
   //-------------HEAD #5 PARAMETERS--------------------------

   "PLANT_CONSTANTS".CONST_rgtHeadPar[4].dParametersToDownload := 17;

   //Parameter IOfunct_LIO1
   "PLANT_CONSTANTS".CONST_rgtHeadPar[4].rgtAxisParameters[0].iAddress := 1826;
   "PLANT_CONSTANTS".CONST_rgtHeadPar[4].rgtAxisParameters[0].iLength := 2;
   "PLANT_CONSTANTS".CONST_rgtHeadPar[4].rgtAxisParameters[0].dValue := 20;

   //Parameter IOfunct_LIO2
   "PLANT_CONSTANTS".CONST_rgtHeadPar[4].rgtAxisParameters[1].iAddress := 1828;
   "PLANT_CONSTANTS".CONST_rgtHeadPar[4].rgtAxisParameters[1].iLength := 2;
   "PLANT_CONSTANTS".CONST_rgtHeadPar[4].rgtAxisParameters[1].dValue := 1;

   //Parameter IOfunct_LIO3
   "PLANT_CONSTANTS".CONST_rgtHeadPar[4].rgtAxisParameters[2].iAddress := 1830;
   "PLANT_CONSTANTS".CONST_rgtHeadPar[4].rgtAxisParameters[2].iLength := 2;
   "PLANT_CONSTANTS".CONST_rgtHeadPar[4].rgtAxisParameters[2].dValue := 1;

   //Parameter IOfunct_LIO4
   "PLANT_CONSTANTS".CONST_rgtHeadPar[4].rgtAxisParameters[3].iAddress := 1832;
   "PLANT_CONSTANTS".CONST_rgtHeadPar[4].rgtAxisParameters[3].iLength := 2;
   "PLANT_CONSTANTS".CONST_rgtHeadPar[4].rgtAxisParameters[3].dValue := 1;

   //Parameter IOsigLimN
   "PLANT_CONSTANTS".CONST_rgtHeadPar[4].rgtAxisParameters[4].iAddress := 1566;
   "PLANT_CONSTANTS".CONST_rgtHeadPar[4].rgtAxisParameters[4].iLength := 2;
   "PLANT_CONSTANTS".CONST_rgtHeadPar[4].rgtAxisParameters[4].dValue := 0;

   //Parameter IOsigLimP
   "PLANT_CONSTANTS".CONST_rgtHeadPar[4].rgtAxisParameters[5].iAddress := 1568;
   "PLANT_CONSTANTS".CONST_rgtHeadPar[4].rgtAxisParameters[5].iLength := 2;
   "PLANT_CONSTANTS".CONST_rgtHeadPar[4].rgtAxisParameters[5].dValue := 0;

   //Parameter IOsigRef
   "PLANT_CONSTANTS".CONST_rgtHeadPar[4].rgtAxisParameters[6].iAddress := 1564;
   "PLANT_CONSTANTS".CONST_rgtHeadPar[4].rgtAxisParameters[6].iLength := 2;
   "PLANT_CONSTANTS".CONST_rgtHeadPar[4].rgtAxisParameters[6].dValue := 2;

   //Parameter POSdirOfRotat
   "PLANT_CONSTANTS".CONST_rgtHeadPar[4].rgtAxisParameters[7].iAddress := 1560;
   "PLANT_CONSTANTS".CONST_rgtHeadPar[4].rgtAxisParameters[7].iLength := 2;
   "PLANT_CONSTANTS".CONST_rgtHeadPar[4].rgtAxisParameters[7].dValue := 0;

   //Parameter POSscaleDenom
   "PLANT_CONSTANTS".CONST_rgtHeadPar[4].rgtAxisParameters[8].iAddress := 1550;
   "PLANT_CONSTANTS".CONST_rgtHeadPar[4].rgtAxisParameters[8].iLength := 4;
   "PLANT_CONSTANTS".CONST_rgtHeadPar[4].rgtAxisParameters[8].dValue := 500;

   //Parameter POSscaleNum
   "PLANT_CONSTANTS".CONST_rgtHeadPar[4].rgtAxisParameters[9].iAddress := 1552;
   "PLANT_CONSTANTS".CONST_rgtHeadPar[4].rgtAxisParameters[9].iLength := 4;
   "PLANT_CONSTANTS".CONST_rgtHeadPar[4].rgtAxisParameters[9].dValue := 1;

   //Parameter RAMPacc
   "PLANT_CONSTANTS".CONST_rgtHeadPar[4].rgtAxisParameters[10].iAddress := 1556;
   "PLANT_CONSTANTS".CONST_rgtHeadPar[4].rgtAxisParameters[10].iLength := 4;
   "PLANT_CONSTANTS".CONST_rgtHeadPar[4].rgtAxisParameters[10].dValue := 20000;//[rot/s2]

   //Parameter RAMPdecel
   "PLANT_CONSTANTS".CONST_rgtHeadPar[4].rgtAxisParameters[11].iAddress := 1558;
   "PLANT_CONSTANTS".CONST_rgtHeadPar[4].rgtAxisParameters[11].iLength := 4;
   "PLANT_CONSTANTS".CONST_rgtHeadPar[4].rgtAxisParameters[11].dValue := 20000;//[rot/s2]

   //Parameter JOGn_fast
   "PLANT_CONSTANTS".CONST_rgtHeadPar[4].rgtAxisParameters[12].iAddress := 10506;
   "PLANT_CONSTANTS".CONST_rgtHeadPar[4].rgtAxisParameters[12].iLength := 2;
   "PLANT_CONSTANTS".CONST_rgtHeadPar[4].rgtAxisParameters[12].dValue := 1000;//[rot/min]

   //Parameter JOGn_slow
   "PLANT_CONSTANTS".CONST_rgtHeadPar[4].rgtAxisParameters[13].iAddress := 10504;
   "PLANT_CONSTANTS".CONST_rgtHeadPar[4].rgtAxisParameters[13].iLength := 2;
   "PLANT_CONSTANTS".CONST_rgtHeadPar[4].rgtAxisParameters[13].dValue := 1000;//[rot/min]

   //Parameter JOGstepusr
   "PLANT_CONSTANTS".CONST_rgtHeadPar[4].rgtAxisParameters[14].iAddress := 10510;
   "PLANT_CONSTANTS".CONST_rgtHeadPar[4].rgtAxisParameters[14].iLength := 4;
   "PLANT_CONSTANTS".CONST_rgtHeadPar[4].rgtAxisParameters[14].dValue := 0;

   //Parameter JOGtime
   "PLANT_CONSTANTS".CONST_rgtHeadPar[4].rgtAxisParameters[15].iAddress := 10512;
   "PLANT_CONSTANTS".CONST_rgtHeadPar[4].rgtAxisParameters[15].iLength := 2;
   "PLANT_CONSTANTS".CONST_rgtHeadPar[4].rgtAxisParameters[15].dValue := 1;

   //Parameter PAReeprSave ---MUST BE THE LAST!!!
   "PLANT_CONSTANTS".CONST_rgtHeadPar[4].rgtAxisParameters[16].iAddress := 1026;
   "PLANT_CONSTANTS".CONST_rgtHeadPar[4].rgtAxisParameters[16].iLength := 2;
   "PLANT_CONSTANTS".CONST_rgtHeadPar[4].rgtAxisParameters[16].dValue := 1;


   //-------------HEAD #6 PARAMETERS--------------------------

   "PLANT_CONSTANTS".CONST_rgtHeadPar[5].dParametersToDownload := 17;

   //Parameter IOfunct_LIO1
   "PLANT_CONSTANTS".CONST_rgtHeadPar[5].rgtAxisParameters[0].iAddress := 1826;
   "PLANT_CONSTANTS".CONST_rgtHeadPar[5].rgtAxisParameters[0].iLength := 2;
   "PLANT_CONSTANTS".CONST_rgtHeadPar[5].rgtAxisParameters[0].dValue := 20;

   //Parameter IOfunct_LIO2
   "PLANT_CONSTANTS".CONST_rgtHeadPar[5].rgtAxisParameters[1].iAddress := 1828;
   "PLANT_CONSTANTS".CONST_rgtHeadPar[5].rgtAxisParameters[1].iLength := 2;
   "PLANT_CONSTANTS".CONST_rgtHeadPar[5].rgtAxisParameters[1].dValue := 1;

   //Parameter IOfunct_LIO3
   "PLANT_CONSTANTS".CONST_rgtHeadPar[5].rgtAxisParameters[2].iAddress := 1830;
   "PLANT_CONSTANTS".CONST_rgtHeadPar[5].rgtAxisParameters[2].iLength := 2;
   "PLANT_CONSTANTS".CONST_rgtHeadPar[5].rgtAxisParameters[2].dValue := 1;

   //Parameter IOfunct_LIO4
   "PLANT_CONSTANTS".CONST_rgtHeadPar[5].rgtAxisParameters[3].iAddress := 1832;
   "PLANT_CONSTANTS".CONST_rgtHeadPar[5].rgtAxisParameters[3].iLength := 2;
   "PLANT_CONSTANTS".CONST_rgtHeadPar[5].rgtAxisParameters[3].dValue := 1;

   //Parameter IOsigLimN
   "PLANT_CONSTANTS".CONST_rgtHeadPar[5].rgtAxisParameters[4].iAddress := 1566;
   "PLANT_CONSTANTS".CONST_rgtHeadPar[5].rgtAxisParameters[4].iLength := 2;
   "PLANT_CONSTANTS".CONST_rgtHeadPar[5].rgtAxisParameters[4].dValue := 0;

   //Parameter IOsigLimP
   "PLANT_CONSTANTS".CONST_rgtHeadPar[5].rgtAxisParameters[5].iAddress := 1568;
   "PLANT_CONSTANTS".CONST_rgtHeadPar[5].rgtAxisParameters[5].iLength := 2;
   "PLANT_CONSTANTS".CONST_rgtHeadPar[5].rgtAxisParameters[5].dValue := 0;

   //Parameter IOsigRef
   "PLANT_CONSTANTS".CONST_rgtHeadPar[5].rgtAxisParameters[6].iAddress := 1564;
   "PLANT_CONSTANTS".CONST_rgtHeadPar[5].rgtAxisParameters[6].iLength := 2;
   "PLANT_CONSTANTS".CONST_rgtHeadPar[5].rgtAxisParameters[6].dValue := 2;

   //Parameter POSdirOfRotat
   "PLANT_CONSTANTS".CONST_rgtHeadPar[5].rgtAxisParameters[7].iAddress := 1560;
   "PLANT_CONSTANTS".CONST_rgtHeadPar[5].rgtAxisParameters[7].iLength := 2;
   "PLANT_CONSTANTS".CONST_rgtHeadPar[5].rgtAxisParameters[7].dValue := 0;

   //Parameter POSscaleDenom
   "PLANT_CONSTANTS".CONST_rgtHeadPar[5].rgtAxisParameters[8].iAddress := 1550;
   "PLANT_CONSTANTS".CONST_rgtHeadPar[5].rgtAxisParameters[8].iLength := 4;
   "PLANT_CONSTANTS".CONST_rgtHeadPar[5].rgtAxisParameters[8].dValue := 500;

   //Parameter POSscaleNum
   "PLANT_CONSTANTS".CONST_rgtHeadPar[5].rgtAxisParameters[9].iAddress := 1552;
   "PLANT_CONSTANTS".CONST_rgtHeadPar[5].rgtAxisParameters[9].iLength := 4;
   "PLANT_CONSTANTS".CONST_rgtHeadPar[5].rgtAxisParameters[9].dValue := 1;

   //Parameter RAMPacc
   "PLANT_CONSTANTS".CONST_rgtHeadPar[5].rgtAxisParameters[10].iAddress := 1556;
   "PLANT_CONSTANTS".CONST_rgtHeadPar[5].rgtAxisParameters[10].iLength := 4;
   "PLANT_CONSTANTS".CONST_rgtHeadPar[5].rgtAxisParameters[10].dValue := 20000;//[rot/s2]

   //Parameter RAMPdecel
   "PLANT_CONSTANTS".CONST_rgtHeadPar[5].rgtAxisParameters[11].iAddress := 1558;
   "PLANT_CONSTANTS".CONST_rgtHeadPar[5].rgtAxisParameters[11].iLength := 4;
   "PLANT_CONSTANTS".CONST_rgtHeadPar[5].rgtAxisParameters[11].dValue := 20000;//[rot/s2]

   //Parameter JOGn_fast
   "PLANT_CONSTANTS".CONST_rgtHeadPar[5].rgtAxisParameters[12].iAddress := 10506;
   "PLANT_CONSTANTS".CONST_rgtHeadPar[5].rgtAxisParameters[12].iLength := 2;
   "PLANT_CONSTANTS".CONST_rgtHeadPar[5].rgtAxisParameters[12].dValue := 1000;//[rot/min]

   //Parameter JOGn_slow
   "PLANT_CONSTANTS".CONST_rgtHeadPar[5].rgtAxisParameters[13].iAddress := 10504;
   "PLANT_CONSTANTS".CONST_rgtHeadPar[5].rgtAxisParameters[13].iLength := 2;
   "PLANT_CONSTANTS".CONST_rgtHeadPar[5].rgtAxisParameters[13].dValue := 1000;//[rot/min]

   //Parameter JOGstepusr
   "PLANT_CONSTANTS".CONST_rgtHeadPar[5].rgtAxisParameters[14].iAddress := 10510;
   "PLANT_CONSTANTS".CONST_rgtHeadPar[5].rgtAxisParameters[14].iLength := 4;
   "PLANT_CONSTANTS".CONST_rgtHeadPar[5].rgtAxisParameters[14].dValue := 0;

   //Parameter JOGtime
   "PLANT_CONSTANTS".CONST_rgtHeadPar[5].rgtAxisParameters[15].iAddress := 10512;
   "PLANT_CONSTANTS".CONST_rgtHeadPar[5].rgtAxisParameters[15].iLength := 2;
   "PLANT_CONSTANTS".CONST_rgtHeadPar[5].rgtAxisParameters[15].dValue := 1;

   //Parameter PAReeprSave ---MUST BE THE LAST!!!
   "PLANT_CONSTANTS".CONST_rgtHeadPar[5].rgtAxisParameters[16].iAddress := 1026;
   "PLANT_CONSTANTS".CONST_rgtHeadPar[5].rgtAxisParameters[16].iLength := 2;
   "PLANT_CONSTANTS".CONST_rgtHeadPar[5].rgtAxisParameters[16].dValue := 1;


   //-------------HEAD #6 PARAMETERS--------------------------

   "PLANT_CONSTANTS".CONST_rgtHeadPar[6].dParametersToDownload := 17;

   //Parameter IOfunct_LIO1
   "PLANT_CONSTANTS".CONST_rgtHeadPar[6].rgtAxisParameters[0].iAddress := 1826;
   "PLANT_CONSTANTS".CONST_rgtHeadPar[6].rgtAxisParameters[0].iLength := 2;
   "PLANT_CONSTANTS".CONST_rgtHeadPar[6].rgtAxisParameters[0].dValue := 20;

   //Parameter IOfunct_LIO2
   "PLANT_CONSTANTS".CONST_rgtHeadPar[6].rgtAxisParameters[1].iAddress := 1828;
   "PLANT_CONSTANTS".CONST_rgtHeadPar[6].rgtAxisParameters[1].iLength := 2;
   "PLANT_CONSTANTS".CONST_rgtHeadPar[6].rgtAxisParameters[1].dValue := 1;

   //Parameter IOfunct_LIO3
   "PLANT_CONSTANTS".CONST_rgtHeadPar[6].rgtAxisParameters[2].iAddress := 1830;
   "PLANT_CONSTANTS".CONST_rgtHeadPar[6].rgtAxisParameters[2].iLength := 2;
   "PLANT_CONSTANTS".CONST_rgtHeadPar[6].rgtAxisParameters[2].dValue := 1;

   //Parameter IOfunct_LIO4
   "PLANT_CONSTANTS".CONST_rgtHeadPar[6].rgtAxisParameters[3].iAddress := 1832;
   "PLANT_CONSTANTS".CONST_rgtHeadPar[6].rgtAxisParameters[3].iLength := 2;
   "PLANT_CONSTANTS".CONST_rgtHeadPar[6].rgtAxisParameters[3].dValue := 1;

   //Parameter IOsigLimN
   "PLANT_CONSTANTS".CONST_rgtHeadPar[6].rgtAxisParameters[4].iAddress := 1566;
   "PLANT_CONSTANTS".CONST_rgtHeadPar[6].rgtAxisParameters[4].iLength := 2;
   "PLANT_CONSTANTS".CONST_rgtHeadPar[6].rgtAxisParameters[4].dValue := 0;

   //Parameter IOsigLimP
   "PLANT_CONSTANTS".CONST_rgtHeadPar[6].rgtAxisParameters[5].iAddress := 1568;
   "PLANT_CONSTANTS".CONST_rgtHeadPar[6].rgtAxisParameters[5].iLength := 2;
   "PLANT_CONSTANTS".CONST_rgtHeadPar[6].rgtAxisParameters[5].dValue := 0;

   //Parameter IOsigRef
   "PLANT_CONSTANTS".CONST_rgtHeadPar[6].rgtAxisParameters[6].iAddress := 1564;
   "PLANT_CONSTANTS".CONST_rgtHeadPar[6].rgtAxisParameters[6].iLength := 2;
   "PLANT_CONSTANTS".CONST_rgtHeadPar[6].rgtAxisParameters[6].dValue := 2;

   //Parameter POSdirOfRotat
   "PLANT_CONSTANTS".CONST_rgtHeadPar[6].rgtAxisParameters[7].iAddress := 1560;
   "PLANT_CONSTANTS".CONST_rgtHeadPar[6].rgtAxisParameters[7].iLength := 2;
   "PLANT_CONSTANTS".CONST_rgtHeadPar[6].rgtAxisParameters[7].dValue := 0;

   //Parameter POSscaleDenom
   "PLANT_CONSTANTS".CONST_rgtHeadPar[6].rgtAxisParameters[8].iAddress := 1550;
   "PLANT_CONSTANTS".CONST_rgtHeadPar[6].rgtAxisParameters[8].iLength := 4;
   "PLANT_CONSTANTS".CONST_rgtHeadPar[6].rgtAxisParameters[8].dValue := 500;

   //Parameter POSscaleNum
   "PLANT_CONSTANTS".CONST_rgtHeadPar[6].rgtAxisParameters[9].iAddress := 1552;
   "PLANT_CONSTANTS".CONST_rgtHeadPar[6].rgtAxisParameters[9].iLength := 4;
   "PLANT_CONSTANTS".CONST_rgtHeadPar[6].rgtAxisParameters[9].dValue := 1;

   //Parameter RAMPacc
   "PLANT_CONSTANTS".CONST_rgtHeadPar[6].rgtAxisParameters[10].iAddress := 1556;
   "PLANT_CONSTANTS".CONST_rgtHeadPar[6].rgtAxisParameters[10].iLength := 4;
   "PLANT_CONSTANTS".CONST_rgtHeadPar[6].rgtAxisParameters[10].dValue := 20000;//[rot/s2]

   //Parameter RAMPdecel
   "PLANT_CONSTANTS".CONST_rgtHeadPar[6].rgtAxisParameters[11].iAddress := 1558;
   "PLANT_CONSTANTS".CONST_rgtHeadPar[6].rgtAxisParameters[11].iLength := 4;
   "PLANT_CONSTANTS".CONST_rgtHeadPar[6].rgtAxisParameters[11].dValue := 20000;//[rot/s2]

   //Parameter JOGn_fast
   "PLANT_CONSTANTS".CONST_rgtHeadPar[6].rgtAxisParameters[12].iAddress := 10506;
   "PLANT_CONSTANTS".CONST_rgtHeadPar[6].rgtAxisParameters[12].iLength := 2;
   "PLANT_CONSTANTS".CONST_rgtHeadPar[6].rgtAxisParameters[12].dValue := 1000;//[rot/min]

   //Parameter JOGn_slow
   "PLANT_CONSTANTS".CONST_rgtHeadPar[6].rgtAxisParameters[13].iAddress := 10504;
   "PLANT_CONSTANTS".CONST_rgtHeadPar[6].rgtAxisParameters[13].iLength := 2;
   "PLANT_CONSTANTS".CONST_rgtHeadPar[6].rgtAxisParameters[13].dValue := 1000;//[rot/min]

   //Parameter JOGstepusr
   "PLANT_CONSTANTS".CONST_rgtHeadPar[6].rgtAxisParameters[14].iAddress := 10510;
   "PLANT_CONSTANTS".CONST_rgtHeadPar[6].rgtAxisParameters[14].iLength := 4;
   "PLANT_CONSTANTS".CONST_rgtHeadPar[6].rgtAxisParameters[14].dValue := 0;

   //Parameter JOGtime
   "PLANT_CONSTANTS".CONST_rgtHeadPar[6].rgtAxisParameters[15].iAddress := 10512;
   "PLANT_CONSTANTS".CONST_rgtHeadPar[6].rgtAxisParameters[15].iLength := 2;
   "PLANT_CONSTANTS".CONST_rgtHeadPar[6].rgtAxisParameters[15].dValue := 1;

   //Parameter PAReeprSave ---MUST BE THE LAST!!!
   "PLANT_CONSTANTS".CONST_rgtHeadPar[6].rgtAxisParameters[16].iAddress := 1026;
   "PLANT_CONSTANTS".CONST_rgtHeadPar[6].rgtAxisParameters[16].iLength := 2;
   "PLANT_CONSTANTS".CONST_rgtHeadPar[6].rgtAxisParameters[16].dValue := 1;


   //-------------HEAD #8 PARAMETERS--------------------------

   "PLANT_CONSTANTS".CONST_rgtHeadPar[7].dParametersToDownload := 17;

   //Parameter IOfunct_LIO1
   "PLANT_CONSTANTS".CONST_rgtHeadPar[7].rgtAxisParameters[0].iAddress := 1826;
   "PLANT_CONSTANTS".CONST_rgtHeadPar[7].rgtAxisParameters[0].iLength := 2;
   "PLANT_CONSTANTS".CONST_rgtHeadPar[7].rgtAxisParameters[0].dValue := 20;

   //Parameter IOfunct_LIO2
   "PLANT_CONSTANTS".CONST_rgtHeadPar[7].rgtAxisParameters[1].iAddress := 1828;
   "PLANT_CONSTANTS".CONST_rgtHeadPar[7].rgtAxisParameters[1].iLength := 2;
   "PLANT_CONSTANTS".CONST_rgtHeadPar[7].rgtAxisParameters[1].dValue := 1;

   //Parameter IOfunct_LIO3
   "PLANT_CONSTANTS".CONST_rgtHeadPar[7].rgtAxisParameters[2].iAddress := 1830;
   "PLANT_CONSTANTS".CONST_rgtHeadPar[7].rgtAxisParameters[2].iLength := 2;
   "PLANT_CONSTANTS".CONST_rgtHeadPar[7].rgtAxisParameters[2].dValue := 1;

   //Parameter IOfunct_LIO4
   "PLANT_CONSTANTS".CONST_rgtHeadPar[7].rgtAxisParameters[3].iAddress := 1832;
   "PLANT_CONSTANTS".CONST_rgtHeadPar[7].rgtAxisParameters[3].iLength := 2;
   "PLANT_CONSTANTS".CONST_rgtHeadPar[7].rgtAxisParameters[3].dValue := 1;

   //Parameter IOsigLimN
   "PLANT_CONSTANTS".CONST_rgtHeadPar[7].rgtAxisParameters[4].iAddress := 1566;
   "PLANT_CONSTANTS".CONST_rgtHeadPar[7].rgtAxisParameters[4].iLength := 2;
   "PLANT_CONSTANTS".CONST_rgtHeadPar[7].rgtAxisParameters[4].dValue := 0;

   //Parameter IOsigLimP
   "PLANT_CONSTANTS".CONST_rgtHeadPar[7].rgtAxisParameters[5].iAddress := 1568;
   "PLANT_CONSTANTS".CONST_rgtHeadPar[7].rgtAxisParameters[5].iLength := 2;
   "PLANT_CONSTANTS".CONST_rgtHeadPar[7].rgtAxisParameters[5].dValue := 0;

   //Parameter IOsigRef
   "PLANT_CONSTANTS".CONST_rgtHeadPar[7].rgtAxisParameters[6].iAddress := 1564;
   "PLANT_CONSTANTS".CONST_rgtHeadPar[7].rgtAxisParameters[6].iLength := 2;
   "PLANT_CONSTANTS".CONST_rgtHeadPar[7].rgtAxisParameters[6].dValue := 2;

   //Parameter POSdirOfRotat
   "PLANT_CONSTANTS".CONST_rgtHeadPar[7].rgtAxisParameters[7].iAddress := 1560;
   "PLANT_CONSTANTS".CONST_rgtHeadPar[7].rgtAxisParameters[7].iLength := 2;
   "PLANT_CONSTANTS".CONST_rgtHeadPar[7].rgtAxisParameters[7].dValue := 0;

   //Parameter POSscaleDenom
   "PLANT_CONSTANTS".CONST_rgtHeadPar[7].rgtAxisParameters[8].iAddress := 1550;
   "PLANT_CONSTANTS".CONST_rgtHeadPar[7].rgtAxisParameters[8].iLength := 4;
   "PLANT_CONSTANTS".CONST_rgtHeadPar[7].rgtAxisParameters[8].dValue := 500;

   //Parameter POSscaleNum
   "PLANT_CONSTANTS".CONST_rgtHeadPar[7].rgtAxisParameters[9].iAddress := 1552;
   "PLANT_CONSTANTS".CONST_rgtHeadPar[7].rgtAxisParameters[9].iLength := 4;
   "PLANT_CONSTANTS".CONST_rgtHeadPar[7].rgtAxisParameters[9].dValue := 1;

   //Parameter RAMPacc
   "PLANT_CONSTANTS".CONST_rgtHeadPar[7].rgtAxisParameters[10].iAddress := 1556;
   "PLANT_CONSTANTS".CONST_rgtHeadPar[7].rgtAxisParameters[10].iLength := 4;
   "PLANT_CONSTANTS".CONST_rgtHeadPar[7].rgtAxisParameters[10].dValue := 20000;//[rot/s2]

   //Parameter RAMPdecel
   "PLANT_CONSTANTS".CONST_rgtHeadPar[7].rgtAxisParameters[11].iAddress := 1558;
   "PLANT_CONSTANTS".CONST_rgtHeadPar[7].rgtAxisParameters[11].iLength := 4;
   "PLANT_CONSTANTS".CONST_rgtHeadPar[7].rgtAxisParameters[11].dValue := 20000;//[rot/s2]

   //Parameter JOGn_fast
   "PLANT_CONSTANTS".CONST_rgtHeadPar[7].rgtAxisParameters[12].iAddress := 10506;
   "PLANT_CONSTANTS".CONST_rgtHeadPar[7].rgtAxisParameters[12].iLength := 2;
   "PLANT_CONSTANTS".CONST_rgtHeadPar[7].rgtAxisParameters[12].dValue := 1000;//[rot/min]

   //Parameter JOGn_slow
   "PLANT_CONSTANTS".CONST_rgtHeadPar[7].rgtAxisParameters[13].iAddress := 10504;
   "PLANT_CONSTANTS".CONST_rgtHeadPar[7].rgtAxisParameters[13].iLength := 2;
   "PLANT_CONSTANTS".CONST_rgtHeadPar[7].rgtAxisParameters[13].dValue := 1000;//[rot/min]

   //Parameter JOGstepusr
   "PLANT_CONSTANTS".CONST_rgtHeadPar[7].rgtAxisParameters[14].iAddress := 10510;
   "PLANT_CONSTANTS".CONST_rgtHeadPar[7].rgtAxisParameters[14].iLength := 4;
   "PLANT_CONSTANTS".CONST_rgtHeadPar[7].rgtAxisParameters[14].dValue := 0;

   //Parameter JOGtime
   "PLANT_CONSTANTS".CONST_rgtHeadPar[7].rgtAxisParameters[15].iAddress := 10512;
   "PLANT_CONSTANTS".CONST_rgtHeadPar[7].rgtAxisParameters[15].iLength := 2;
   "PLANT_CONSTANTS".CONST_rgtHeadPar[7].rgtAxisParameters[15].dValue := 1;

   //Parameter PAReeprSave ---MUST BE THE LAST!!!
   "PLANT_CONSTANTS".CONST_rgtHeadPar[7].rgtAxisParameters[16].iAddress := 1026;
   "PLANT_CONSTANTS".CONST_rgtHeadPar[7].rgtAxisParameters[16].iLength := 2;
   "PLANT_CONSTANTS".CONST_rgtHeadPar[7].rgtAxisParameters[16].dValue := 1;





   //Home position #Head 1
   "M256_Manag_IDB".M256M_IDB[0].ILx2T_Homing_Instance.i_inHM_method := 11;
   "M256_Manag_IDB".M256M_IDB[0].ILx2T_Homing_Instance.i_inHMn:= 500;
   "M256_Manag_IDB".M256M_IDB[0].ILx2T_Homing_Instance.i_inHMn_out := 10;
   "M256_Manag_IDB".M256M_IDB[0].ILx2T_Homing_Instance.i_diHMoutdisusr:= 0;
   "M256_Manag_IDB".M256M_IDB[0].ILx2T_Homing_Instance.i_diHMdisusr:= 1;

   //Home position #Head 2
   "M256_Manag_IDB".M256M_IDB[1].ILx2T_Homing_Instance.i_inHM_method := 11;
   "M256_Manag_IDB".M256M_IDB[1].ILx2T_Homing_Instance.i_inHMn := 500;
   "M256_Manag_IDB".M256M_IDB[1].ILx2T_Homing_Instance.i_inHMn_out := 10;
   "M256_Manag_IDB".M256M_IDB[1].ILx2T_Homing_Instance.i_diHMoutdisusr:= 0;
   "M256_Manag_IDB".M256M_IDB[1].ILx2T_Homing_Instance.i_diHMdisusr:= 1;

   //Home position #Head 3
   "M256_Manag_IDB".M256M_IDB[2].ILx2T_Homing_Instance.i_inHM_method := 11;
   "M256_Manag_IDB".M256M_IDB[2].ILx2T_Homing_Instance.i_inHMn := 500;
   "M256_Manag_IDB".M256M_IDB[2].ILx2T_Homing_Instance.i_inHMn_out := 10;
   "M256_Manag_IDB".M256M_IDB[2].ILx2T_Homing_Instance.i_diHMoutdisusr:= 0;
   "M256_Manag_IDB".M256M_IDB[2].ILx2T_Homing_Instance.i_diHMdisusr:= 1;

   //Home position #Head 4
   "M256_Manag_IDB".M256M_IDB[3].ILx2T_Homing_Instance.i_inHM_method := 11;
   "M256_Manag_IDB".M256M_IDB[3].ILx2T_Homing_Instance.i_inHMn := 500;
   "M256_Manag_IDB".M256M_IDB[3].ILx2T_Homing_Instance.i_inHMn_out := 10;
   "M256_Manag_IDB".M256M_IDB[3].ILx2T_Homing_Instance.i_diHMoutdisusr:= 0;
   "M256_Manag_IDB".M256M_IDB[3].ILx2T_Homing_Instance.i_diHMdisusr:= 1;

   //Home position #Head 5
   "M256_Manag_IDB".M256M_IDB[4].ILx2T_Homing_Instance.i_inHM_method := 7;
   "M256_Manag_IDB".M256M_IDB[4].ILx2T_Homing_Instance.i_inHMn := 500;
   "M256_Manag_IDB".M256M_IDB[4].ILx2T_Homing_Instance.i_inHMn_out := 10;
   "M256_Manag_IDB".M256M_IDB[4].ILx2T_Homing_Instance.i_diHMoutdisusr := 0;
   "M256_Manag_IDB".M256M_IDB[4].ILx2T_Homing_Instance.i_diHMdisusr := 1;

   //Home position #Head 6
   "M256_Manag_IDB".M256M_IDB[5].ILx2T_Homing_Instance.i_inHM_method := 7;
   "M256_Manag_IDB".M256M_IDB[5].ILx2T_Homing_Instance.i_inHMn := 500;
   "M256_Manag_IDB".M256M_IDB[5].ILx2T_Homing_Instance.i_inHMn_out := 10;
   "M256_Manag_IDB".M256M_IDB[5].ILx2T_Homing_Instance.i_diHMoutdisusr := 0;
   "M256_Manag_IDB".M256M_IDB[5].ILx2T_Homing_Instance.i_diHMdisusr := 1;

   //Home position #Head 7
   "M256_Manag_IDB".M256M_IDB[6].ILx2T_Homing_Instance.i_inHM_method := 7;
   "M256_Manag_IDB".M256M_IDB[6].ILx2T_Homing_Instance.i_inHMn := 500;
   "M256_Manag_IDB".M256M_IDB[6].ILx2T_Homing_Instance.i_inHMn_out := 10;
   "M256_Manag_IDB".M256M_IDB[6].ILx2T_Homing_Instance.i_diHMoutdisusr := 0;
   "M256_Manag_IDB".M256M_IDB[6].ILx2T_Homing_Instance.i_diHMdisusr := 1;

   //Home position #Head 8
   "M256_Manag_IDB".M256M_IDB[7].ILx2T_Homing_Instance.i_inHM_method := 7;
   "M256_Manag_IDB".M256M_IDB[7].ILx2T_Homing_Instance.i_inHMn := 500;
   "M256_Manag_IDB".M256M_IDB[7].ILx2T_Homing_Instance.i_inHMn_out := 10;
   "M256_Manag_IDB".M256M_IDB[7].ILx2T_Homing_Instance.i_diHMoutdisusr := 0;
   "M256_Manag_IDB".M256M_IDB[7].ILx2T_Homing_Instance.i_diHMdisusr := 1;


   //Positioning Head #1
   "M256_Manag_IDB".M256M_IDB[0].ILx2T_ProfilePosition_Instance.i_inTargetVelocity := 4300; 

   //Positioning Head #2
   "M256_Manag_IDB".M256M_IDB[1].ILx2T_ProfilePosition_Instance.i_inTargetVelocity := 4300;

   //Positioning Head #3
   "M256_Manag_IDB".M256M_IDB[2].ILx2T_ProfilePosition_Instance.i_inTargetVelocity:= 4300;

   //Positioning Head #4
   "M256_Manag_IDB".M256M_IDB[3].ILx2T_ProfilePosition_Instance.i_inTargetVelocity := 4300;

   //Positioning Head #5
   "M256_Manag_IDB".M256M_IDB[4].ILx2T_ProfilePosition_Instance.i_inTargetVelocity := 4300;

   //Positioning Head #6
   "M256_Manag_IDB".M256M_IDB[5].ILx2T_ProfilePosition_Instance.i_inTargetVelocity := 4300;

   //Positioning Head #7
   "M256_Manag_IDB".M256M_IDB[6].ILx2T_ProfilePosition_Instance.i_inTargetVelocity := 4300;

   //Positioning Head #8
   "M256_Manag_IDB".M256M_IDB[7].ILx2T_ProfilePosition_Instance.i_inTargetVelocity := 4300;


   //Timeout head initialization
   "M256_Manag_IDB".M256M_IDB[0].AUX_tmHeadInitTimeout.PT := t#20000ms;
   "M256_Manag_IDB".M256M_IDB[1].AUX_tmHeadInitTimeout.PT := t#20000ms;
   "M256_Manag_IDB".M256M_IDB[2].AUX_tmHeadInitTimeout.PT := t#20000ms;
   "M256_Manag_IDB".M256M_IDB[3].AUX_tmHeadInitTimeout.PT := t#20000ms;
   "M256_Manag_IDB".M256M_IDB[4].AUX_tmHeadInitTimeout.PT := t#20000ms;
   "M256_Manag_IDB".M256M_IDB[5].AUX_tmHeadInitTimeout.PT := t#20000ms;
   "M256_Manag_IDB".M256M_IDB[6].AUX_tmHeadInitTimeout.PT := t#20000ms;
   "M256_Manag_IDB".M256M_IDB[7].AUX_tmHeadInitTimeout.PT := t#20000ms;

   //Timeout head homing
   "M256_Manag_IDB".M256M_IDB[0].AUX_tmHeadHomingTimeout.PT := t#60000ms;
   "M256_Manag_IDB".M256M_IDB[1].AUX_tmHeadHomingTimeout.PT := t#60000ms;
   "M256_Manag_IDB".M256M_IDB[2].AUX_tmHeadHomingTimeout.PT := t#60000ms;
   "M256_Manag_IDB".M256M_IDB[3].AUX_tmHeadHomingTimeout.PT := t#60000ms;
   "M256_Manag_IDB".M256M_IDB[4].AUX_tmHeadHomingTimeout.PT := t#60000ms;
   "M256_Manag_IDB".M256M_IDB[5].AUX_tmHeadHomingTimeout.PT := t#60000ms;
   "M256_Manag_IDB".M256M_IDB[6].AUX_tmHeadHomingTimeout.PT := t#60000ms;
   "M256_Manag_IDB".M256M_IDB[7].AUX_tmHeadHomingTimeout.PT := t#60000ms;


   //Timeout head positioning
   "M256_Manag_IDB".M256M_IDB[0].AUX_tmHeadPositioningTimeout.PT := t#6000ms;
   "M256_Manag_IDB".M256M_IDB[1].AUX_tmHeadPositioningTimeout.PT := t#6000ms;
   "M256_Manag_IDB".M256M_IDB[2].AUX_tmHeadPositioningTimeout.PT := t#6000ms;
   "M256_Manag_IDB".M256M_IDB[3].AUX_tmHeadPositioningTimeout.PT := t#6000ms;
   "M256_Manag_IDB".M256M_IDB[4].AUX_tmHeadPositioningTimeout.PT := t#6000ms;
   "M256_Manag_IDB".M256M_IDB[5].AUX_tmHeadPositioningTimeout.PT := t#6000ms;
   "M256_Manag_IDB".M256M_IDB[6].AUX_tmHeadPositioningTimeout.PT := t#6000ms;
   "M256_Manag_IDB".M256M_IDB[7].AUX_tmHeadPositioningTimeout.PT := t#6000ms;


   //Head positioning modality
   "M256_Manag_IDB".M256M_IDB[0].ILx2T_ProfilePosition_Instance.i_inPTP_Type := 1;
   "M256_Manag_IDB".M256M_IDB[1].ILx2T_ProfilePosition_Instance.i_inPTP_Type := 1;
   "M256_Manag_IDB".M256M_IDB[2].ILx2T_ProfilePosition_Instance.i_inPTP_Type := 1;
   "M256_Manag_IDB".M256M_IDB[3].ILx2T_ProfilePosition_Instance.i_inPTP_Type := 1;
   "M256_Manag_IDB".M256M_IDB[4].ILx2T_ProfilePosition_Instance.i_inPTP_Type := 1;
   "M256_Manag_IDB".M256M_IDB[5].ILx2T_ProfilePosition_Instance.i_inPTP_Type := 1;
   "M256_Manag_IDB".M256M_IDB[6].ILx2T_ProfilePosition_Instance.i_inPTP_Type := 1;
   "M256_Manag_IDB".M256M_IDB[7].ILx2T_ProfilePosition_Instance.i_inPTP_Type := 1;
END_FUNCTION

FUNCTION "OUTPUT" : Void   // FC25, LAD
{ S7_Optimized_Access := 'TRUE' }
VERSION : 0.1
   VAR_TEMP
      iRetVal : Int;
      wRetVal : Word;
      xSpareOutput : Bool;
   END_VAR
BEGIN

REGION Network 1 (SCL): Counter card
   "o.1B160AP1.Open_SW_Gate" := "Encoder".OUTPUT_xCounterEnable;
   "o.1B160AP1.Enable_Measure" := "Encoder".OUTPUT_xCounterEnable AND NOT"Encoder".INPUT_xResetEventAcknowledge;
   "o.1B160AP1.Res_Event" :="Encoder".OUTPUT_xResetMeterPulse;
   "o.1B160AP1.CounterCardStatus":P := "o.1B160AP1.CounterCardStatus";
END_REGION

REGION Network 2 (SCL): Cut pressure
   "o.1B160AP1.M217CutPressureHead1":=  "M256_Manag_IDB".M256F_IDB[0].OUTPUT_iPressuremA;
   "o.1B160AP1.M217CutPressureHead2" := "M256_Manag_IDB".M256F_IDB[1].OUTPUT_iPressuremA;
   "o.1B160AP1.M217CutPressureHead3" := "M256_Manag_IDB".M256F_IDB[2].OUTPUT_iPressuremA;
   "o.1B160AP1.M217CutPressureHead4" := "M256_Manag_IDB".M256F_IDB[3].OUTPUT_iPressuremA;
   "o.1B160AP1.M217CutPressureHead5" := "M256_Manag_IDB".M256F_IDB[4].OUTPUT_iPressuremA;
   "o.1B160AP1.M217CutPressureHead6" := "M256_Manag_IDB".M256F_IDB[5].OUTPUT_iPressuremA;
   "o.1B160AP1.M217CutPressureHead7" := "M256_Manag_IDB".M256F_IDB[6].OUTPUT_iPressuremA;
   "o.1B160AP1.M217CutPressureHead8" := "M256_Manag_IDB".M256F_IDB[7].OUTPUT_iPressuremA;
END_REGION

REGION Network 3 (SCL): 151K8
   "o.1B160AP1.1B251HL1.AreaFailure" := "Z256".OUTPUT_xAreaFailure;
   "o.1B160AP1.1B251KA1.ResetLocalEmergency" := "Z256".OUTPUT_xResetLocalEmergency;
END_REGION

REGION Network 4 (SCL): 300A1 / Traffic lighter Lamp
   "o.1B160AP1.M217B1HL5.MachineToMaintenance":= "Z256".OUTPUT_xMachineToMaintenance;
   "o.1B160AP1.M217B1HL6.MachineOutOfOrder":= "Z256".OUTPUT_xMachineOutOfOrder;
   "o.1B160AP1.M217B1HL4.MachineInOrder":= "Z256".OUTPUT_xMachineInOrder;
   "o.1B160AP1.M217B1HL3.MachineReady" :="Z256".OUTPUT_xMachineInOrder;
END_REGION

REGION Network 5 (SCL): Head #1
   "o.1B411AP1.1B411YV2.Head1.CuttingLubrication" :="M256_Manag_IDB".M256F_IDB[0].OUTPUT_xOilON;
   "o.1B411AP1.1B411YV1.Head1.CuttingHeadGlassApproach":="M256_Manag_IDB".M256A_IDB[0].OUTPUT_xCarriageDescent;
   "o.1B411AP1.1B411SA2.Head1.ProductionON" := "Z256".OUTPUT_rgxHeadsInProduction[0];
END_REGION

REGION Network 6 (SCL): Head #2
   "o.1B412AP1.1B412YV2.Head2.CuttingLubrication" := "M256_Manag_IDB".M256F_IDB[1].OUTPUT_xOilON;
   "o.1B412AP1.1B412YV1.Head2.CuttingHeadGlassApproach" := "M256_Manag_IDB".M256A_IDB[1].OUTPUT_xCarriageDescent;
   "o.1B412AP1.1B412SA2.Head2.ProductionON" :="Z256".OUTPUT_rgxHeadsInProduction[1];
END_REGION

REGION Network 7 (SCL): Head #3
   "o.1B413AP1.1B413YV2.Head3.CuttingLubrication" := "M256_Manag_IDB".M256F_IDB[2].OUTPUT_xOilON;
   "o.1B413AP1.1B413YV1.Head3.CuttingHeadGlassApproach":= "M256_Manag_IDB".M256A_IDB[2].OUTPUT_xCarriageDescent;
   "o.1B413AP1.1B413SA2.Head3.ProductionON" := "Z256".OUTPUT_rgxHeadsInProduction[2];
END_REGION

REGION Network 8 (SCL): Head #4
   "o.1B414AP1.1B414YV2.Head4.CuttingLubrication" := "M256_Manag_IDB".M256F_IDB[3].OUTPUT_xOilON;
   "o.1B414AP1.1B414YV1.Head4.CuttingHeadGlassApproach" := "M256_Manag_IDB".M256A_IDB[3].OUTPUT_xCarriageDescent;
   "o.1B414AP1.1B414SA2.Head4.ProductionON":="Z256".OUTPUT_rgxHeadsInProduction[3];
END_REGION

REGION Network 9 (SCL): Head #5
   "o.1B415AP1.1B415YV2.Head5.CuttingLubrication"  := "M256_Manag_IDB".M256F_IDB[4].OUTPUT_xOilON;
   "o.1B415AP1.1B415YV1.Head5.CuttingHeadGlassApproach":="M256_Manag_IDB".M256A_IDB[4].OUTPUT_xCarriageDescent;
   "o.1B415AP1.1B415SA2.Head5.ProductionON" :="Z256".OUTPUT_rgxHeadsInProduction[4];
END_REGION

REGION Network 10 (SCL): Head #6 / Head #5
   "o.1B416AP1.1B416YV2.Head6.CuttingLubrication"  := "M256_Manag_IDB".M256F_IDB[5].OUTPUT_xOilON;
   "o.1B416AP1.1B416YV1.Head6.CuttingHeadGlassApproach":="M256_Manag_IDB".M256A_IDB[5].OUTPUT_xCarriageDescent;
   "o.1B416AP1.1B416SA2.Head6.ProductionON" :="Z256".OUTPUT_rgxHeadsInProduction[5];
END_REGION

REGION Network 11 (SCL): Head #7 / Head #5
   "o.1B417AP1.1B417YV2.Head7.CuttingLubrication"  := "M256_Manag_IDB".M256F_IDB[6].OUTPUT_xOilON;
   "o.1B417AP1.1B417YV1.Head7.CuttingHeadGlassApproach":="M256_Manag_IDB".M256A_IDB[6].OUTPUT_xCarriageDescent;
   "o.1B417AP1.1B417SA2.Head7.ProductionON" := "Z256".OUTPUT_rgxHeadsInProduction[6];
END_REGION

REGION Network 12 (SCL): Head #8 / Head #5
   "o.1B418AP1.1B418YV2.Head8.CuttingLubrication"  := "M256_Manag_IDB".M256F_IDB[7].OUTPUT_xOilON;
   "o.1B418AP1.1B418YV1.Head8.CuttingHeadGlassApproach":="M256_Manag_IDB".M256A_IDB[7].OUTPUT_xCarriageDescent;
   "o.1B418AP1.1B418SA2.Head8.ProductionON" := "Z256".OUTPUT_rgxHeadsInProduction[7];
END_REGION

REGION Network 13 (SCL): Idevice
   "o.IDeviceCPU0" := "CM_IDEV_ToMainLine";
END_REGION
END_FUNCTION

ORGANIZATION_BLOCK "Main"   // OB1, LAD, ProgramCycle
TITLE = "Main Program Sweep (Cycle)"
{ S7_Optimized_Access := 'TRUE' }
VERSION : 0.1
   VAR_INPUT
      Initial_Call : Bool;   // Initial call of this OB
      Remanence : Bool;   // =True, if remanent data are available
   END_VAR
   VAR_TEMP
      TMP_iRetVal : Int;
   END_VAR
   VAR_TEMP   // added for the SCL form of the ladder/FBD networks
      _w1 : Bool;
   END_VAR
BEGIN

REGION Network 1 (SCL): Main

   "OB_Initialize"(FALSE);

   "INPUT"();

   "Encoder_Manager"();

   "Z256_Logic"();



   "CM_Management"();

   "M256_Manag_IDB"();

   "Z256_Output"();

   "SCADA_Mapping"();

   "OUTPUT"();
END_REGION

REGION Network 2: OS gate open
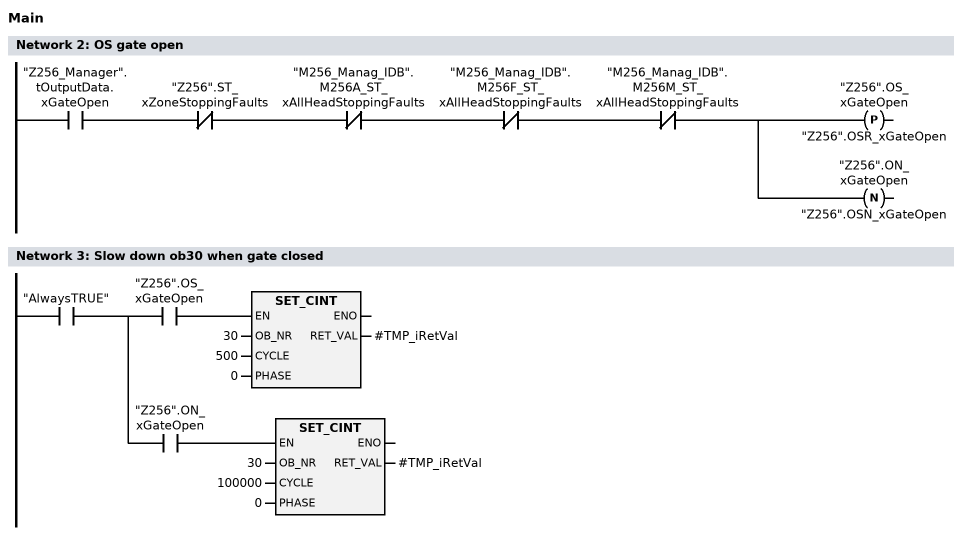
   #_w1 := "Z256_Manager".tOutputData.xGateOpen AND NOT "Z256".ST_xZoneStoppingFaults AND NOT "M256_Manag_IDB".M256A_ST_xAllHeadStoppingFaults AND NOT "M256_Manag_IDB".M256F_ST_xAllHeadStoppingFaults AND NOT "M256_Manag_IDB".M256M_ST_xAllHeadStoppingFaults;
   "Z256".OS_xGateOpen := #_w1 AND NOT "Z256".OSR_xGateOpen;   // rising edge
   "Z256".OSR_xGateOpen := #_w1;
   "Z256".ON_xGateOpen := NOT #_w1 AND "Z256".OSN_xGateOpen;   // falling edge
   "Z256".OSN_xGateOpen := #_w1;
END_REGION

REGION Network 3: Slow down ob30 when gate closed
   #_w1 := "AlwaysTRUE";
   IF "AlwaysTRUE" AND "Z256".OS_xGateOpen THEN
       #TMP_iRetVal := SET_CINT(OB_NR := 30, CYCLE := 500, PHASE := 0);
   END_IF;
   IF #_w1 AND "Z256".ON_xGateOpen THEN
       #TMP_iRetVal := SET_CINT(OB_NR := 30, CYCLE := 100000, PHASE := 0);
   END_IF;
END_REGION
END_ORGANIZATION_BLOCK

ORGANIZATION_BLOCK "Cyclic interrupt"   // OB30, LAD, CyclicInterrupt
{ S7_Optimized_Access := 'TRUE' }
VERSION : 0.1
   VAR_INPUT
      Initial_Call : Bool;   // Initial call of this OB
      Event_Count : Int;   // Events discarded
   END_VAR
   VAR_TEMP
      TMP_dEncValueFast : DInt;
      TMP_xChangeFAST : Bool;
      TMP_dIndexFAST_2 : DInt;
      TMP_dIndexFAST : DInt;
      TMP_dEncoderOverFAST_cmm : DInt;
      TMP_xDummy : Bool;
      TMP_iRetVal : Int;
      TMP_xPressureIncrease : Bool;
   END_VAR
BEGIN

REGION Network 1 (SCL)
   //*************** TASK FAST *************** //
   //Manage the firing  
   IF "CM_Manager".ST_MutingFiringOB = 0 AND "Z256_Manager".tOutputData.xGateOpen THEN

       #TMP_xDummy := false;
       FOR #TMP_dIndexFAST := 0 TO "CONST_dNumberOfHeadsCycle" DO
           IF "Z256_Manager".tOutputData.rgxDataToProcessInter[#TMP_dIndexFAST] <> 0 THEN
               #TMP_xDummy := true;
           END_IF;
       END_FOR;

       IF NOT (#TMP_xDummy) THEN
           RETURN;
       END_IF;

       #TMP_dEncValueFast := DWORD_TO_DINT("i.1B160AP1.CounterActualValue");
       //        #TMP_dEncValueFast := "Encoder".INPUT_dEncoderCounter_count;

       #TMP_xChangeFAST := 0;

       FOR #TMP_dIndexFAST := 0 TO "CONST_dNumberOfHeadsCycle" DO